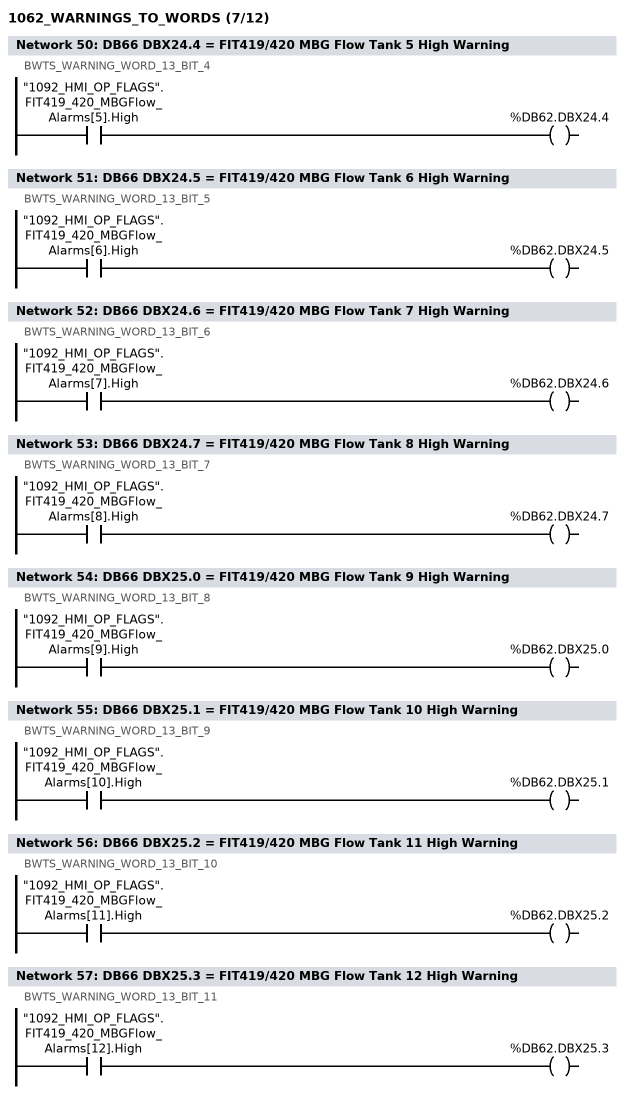
   RUNG wire#powerrail
      Contact( "1092_HMI_OP_FLAGS".FIT419_420_MBGFlow_Alarms[5].High )
      Coil( %DB62.DBX24.4 )
   END_RUNG
   // the same network as SCL:
   %DB62.DBX24.4 := "1092_HMI_OP_FLAGS".FIT419_420_MBGFlow_Alarms[5].High;
END_REGION

REGION Network 51: DB66 DBX24.5 = FIT419/420 MBG Flow Tank 6 High Warning
   // BWTS_WARNING_WORD_13_BIT_5
   RUNG wire#powerrail
      Contact( "1092_HMI_OP_FLAGS".FIT419_420_MBGFlow_Alarms[6].High )
      Coil( %DB62.DBX24.5 )
   END_RUNG
   // the same network as SCL:
   %DB62.DBX24.5 := "1092_HMI_OP_FLAGS".FIT419_420_MBGFlow_Alarms[6].High;
END_REGION

REGION Network 52: DB66 DBX24.6 = FIT419/420 MBG Flow Tank 7 High Warning
   // BWTS_WARNING_WORD_13_BIT_6
   RUNG wire#powerrail
      Contact( "1092_HMI_OP_FLAGS".FIT419_420_MBGFlow_Alarms[7].High )
      Coil( %DB62.DBX24.6 )
   END_RUNG
   // the same network as SCL:
   %DB62.DBX24.6 := "1092_HMI_OP_FLAGS".FIT419_420_MBGFlow_Alarms[7].High;
END_REGION

REGION Network 53: DB66 DBX24.7 = FIT419/420 MBG Flow Tank 8 High Warning
   // BWTS_WARNING_WORD_13_BIT_7
   RUNG wire#powerrail
      Contact( "1092_HMI_OP_FLAGS".FIT419_420_MBGFlow_Alarms[8].High )
      Coil( %DB62.DBX24.7 )
   END_RUNG
   // the same network as SCL:
   %DB62.DBX24.7 := "1092_HMI_OP_FLAGS".FIT419_420_MBGFlow_Alarms[8].High;
END_REGION

REGION Network 54: DB66 DBX25.0 = FIT419/420 MBG Flow Tank 9 High Warning
   // BWTS_WARNING_WORD_13_BIT_8
   RUNG wire#powerrail
      Contact( "1092_HMI_OP_FLAGS".FIT419_420_MBGFlow_Alarms[9].High )
      Coil( %DB62.DBX25.0 )
   END_RUNG
   // the same network as SCL:
   %DB62.DBX25.0 := "1092_HMI_OP_FLAGS".FIT419_420_MBGFlow_Alarms[9].High;
END_REGION

REGION Network 55: DB66 DBX25.1 = FIT419/420 MBG Flow Tank 10 High Warning
   // BWTS_WARNING_WORD_13_BIT_9
   RUNG wire#powerrail
      Contact( "1092_HMI_OP_FLAGS".FIT419_420_MBGFlow_Alarms[10].High )
      Coil( %DB62.DBX25.1 )
   END_RUNG
   // the same network as SCL:
   %DB62.DBX25.1 := "1092_HMI_OP_FLAGS".FIT419_420_MBGFlow_Alarms[10].High;
END_REGION

REGION Network 56: DB66 DBX25.2 = FIT419/420 MBG Flow Tank 11 High Warning
   // BWTS_WARNING_WORD_13_BIT_10
   RUNG wire#powerrail
      Contact( "1092_HMI_OP_FLAGS".FIT419_420_MBGFlow_Alarms[11].High )
      Coil( %DB62.DBX25.2 )
   END_RUNG
   // the same network as SCL:
   %DB62.DBX25.2 := "1092_HMI_OP_FLAGS".FIT419_420_MBGFlow_Alarms[11].High;
END_REGION

REGION Network 57: DB66 DBX25.3 = FIT419/420 MBG Flow Tank 12 High Warning
   // BWTS_WARNING_WORD_13_BIT_11
   RUNG wire#powerrail
      Contact( "1092_HMI_OP_FLAGS".FIT419_420_MBGFlow_Alarms[12].High )
      Coil( %DB62.DBX25.3 )
   END_RUNG
   // the same network as SCL:
   %DB62.DBX25.3 := "1092_HMI_OP_FLAGS".FIT419_420_MBGFlow_Alarms[12].High;
END_REGION

REGION Network 58: DB66 DBX25.4 = FIT419/420 MBG Flow Tank 13 High Warning
   // BWTS_WARNING_WORD_13_BIT_12
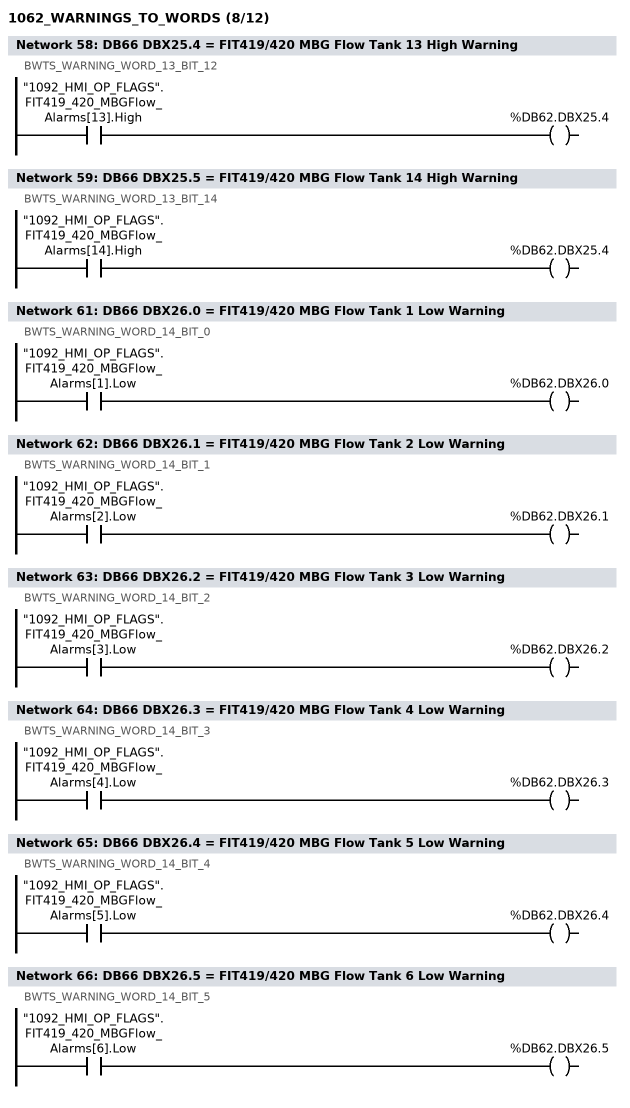
   RUNG wire#powerrail
      Contact( "1092_HMI_OP_FLAGS".FIT419_420_MBGFlow_Alarms[13].High )
      Coil( %DB62.DBX25.4 )
   END_RUNG
   // the same network as SCL:
   %DB62.DBX25.4 := "1092_HMI_OP_FLAGS".FIT419_420_MBGFlow_Alarms[13].High;
END_REGION

REGION Network 59: DB66 DBX25.5 = FIT419/420 MBG Flow Tank 14 High Warning
   // BWTS_WARNING_WORD_13_BIT_14
   RUNG wire#powerrail
      Contact( "1092_HMI_OP_FLAGS".FIT419_420_MBGFlow_Alarms[14].High )
      Coil( %DB62.DBX25.4 )
   END_RUNG
   // the same network as SCL:
   %DB62.DBX25.4 := "1092_HMI_OP_FLAGS".FIT419_420_MBGFlow_Alarms[14].High;
END_REGION

REGION Network 61: DB66 DBX26.0 = FIT419/420 MBG Flow Tank 1 Low Warning
   // BWTS_WARNING_WORD_14_BIT_0
   RUNG wire#powerrail
      Contact( "1092_HMI_OP_FLAGS".FIT419_420_MBGFlow_Alarms[1].Low )
      Coil( %DB62.DBX26.0 )
   END_RUNG
   // the same network as SCL:
   %DB62.DBX26.0 := "1092_HMI_OP_FLAGS".FIT419_420_MBGFlow_Alarms[1].Low;
END_REGION

REGION Network 62: DB66 DBX26.1 = FIT419/420 MBG Flow Tank 2 Low Warning
   // BWTS_WARNING_WORD_14_BIT_1
   RUNG wire#powerrail
      Contact( "1092_HMI_OP_FLAGS".FIT419_420_MBGFlow_Alarms[2].Low )
      Coil( %DB62.DBX26.1 )
   END_RUNG
   // the same network as SCL:
   %DB62.DBX26.1 := "1092_HMI_OP_FLAGS".FIT419_420_MBGFlow_Alarms[2].Low;
END_REGION

REGION Network 63: DB66 DBX26.2 = FIT419/420 MBG Flow Tank 3 Low Warning
   // BWTS_WARNING_WORD_14_BIT_2
   RUNG wire#powerrail
      Contact( "1092_HMI_OP_FLAGS".FIT419_420_MBGFlow_Alarms[3].Low )
      Coil( %DB62.DBX26.2 )
   END_RUNG
   // the same network as SCL:
   %DB62.DBX26.2 := "1092_HMI_OP_FLAGS".FIT419_420_MBGFlow_Alarms[3].Low;
END_REGION

REGION Network 64: DB66 DBX26.3 = FIT419/420 MBG Flow Tank 4 Low Warning
   // BWTS_WARNING_WORD_14_BIT_3
   RUNG wire#powerrail
      Contact( "1092_HMI_OP_FLAGS".FIT419_420_MBGFlow_Alarms[4].Low )
      Coil( %DB62.DBX26.3 )
   END_RUNG
   // the same network as SCL:
   %DB62.DBX26.3 := "1092_HMI_OP_FLAGS".FIT419_420_MBGFlow_Alarms[4].Low;
END_REGION

REGION Network 65: DB66 DBX26.4 = FIT419/420 MBG Flow Tank 5 Low Warning
   // BWTS_WARNING_WORD_14_BIT_4
   RUNG wire#powerrail
      Contact( "1092_HMI_OP_FLAGS".FIT419_420_MBGFlow_Alarms[5].Low )
      Coil( %DB62.DBX26.4 )
   END_RUNG
   // the same network as SCL:
   %DB62.DBX26.4 := "1092_HMI_OP_FLAGS".FIT419_420_MBGFlow_Alarms[5].Low;
END_REGION

REGION Network 66: DB66 DBX26.5 = FIT419/420 MBG Flow Tank 6 Low Warning
   // BWTS_WARNING_WORD_14_BIT_5
   RUNG wire#powerrail
      Contact( "1092_HMI_OP_FLAGS".FIT419_420_MBGFlow_Alarms[6].Low )
      Coil( %DB62.DBX26.5 )
   END_RUNG
   // the same network as SCL:
   %DB62.DBX26.5 := "1092_HMI_OP_FLAGS".FIT419_420_MBGFlow_Alarms[6].Low;
END_REGION

REGION Network 67: DB66 DBX26.6 = FIT419/420 MBG Flow Tank 7 Low Warning
   // BWTS_WARNING_WORD_14_BIT_6
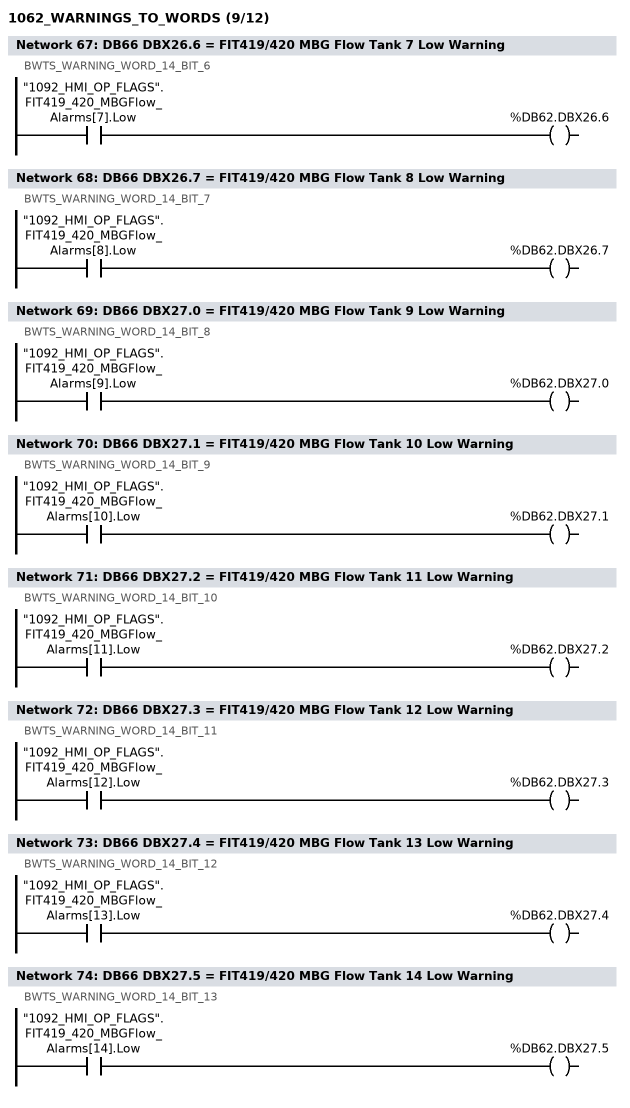
   RUNG wire#powerrail
      Contact( "1092_HMI_OP_FLAGS".FIT419_420_MBGFlow_Alarms[7].Low )
      Coil( %DB62.DBX26.6 )
   END_RUNG
   // the same network as SCL:
   %DB62.DBX26.6 := "1092_HMI_OP_FLAGS".FIT419_420_MBGFlow_Alarms[7].Low;
END_REGION

REGION Network 68: DB66 DBX26.7 = FIT419/420 MBG Flow Tank 8 Low Warning
   // BWTS_WARNING_WORD_14_BIT_7
   RUNG wire#powerrail
      Contact( "1092_HMI_OP_FLAGS".FIT419_420_MBGFlow_Alarms[8].Low )
      Coil( %DB62.DBX26.7 )
   END_RUNG
   // the same network as SCL:
   %DB62.DBX26.7 := "1092_HMI_OP_FLAGS".FIT419_420_MBGFlow_Alarms[8].Low;
END_REGION

REGION Network 69: DB66 DBX27.0 = FIT419/420 MBG Flow Tank 9 Low Warning
   // BWTS_WARNING_WORD_14_BIT_8
   RUNG wire#powerrail
      Contact( "1092_HMI_OP_FLAGS".FIT419_420_MBGFlow_Alarms[9].Low )
      Coil( %DB62.DBX27.0 )
   END_RUNG
   // the same network as SCL:
   %DB62.DBX27.0 := "1092_HMI_OP_FLAGS".FIT419_420_MBGFlow_Alarms[9].Low;
END_REGION

REGION Network 70: DB66 DBX27.1 = FIT419/420 MBG Flow Tank 10 Low Warning
   // BWTS_WARNING_WORD_14_BIT_9
   RUNG wire#powerrail
      Contact( "1092_HMI_OP_FLAGS".FIT419_420_MBGFlow_Alarms[10].Low )
      Coil( %DB62.DBX27.1 )
   END_RUNG
   // the same network as SCL:
   %DB62.DBX27.1 := "1092_HMI_OP_FLAGS".FIT419_420_MBGFlow_Alarms[10].Low;
END_REGION

REGION Network 71: DB66 DBX27.2 = FIT419/420 MBG Flow Tank 11 Low Warning
   // BWTS_WARNING_WORD_14_BIT_10
   RUNG wire#powerrail
      Contact( "1092_HMI_OP_FLAGS".FIT419_420_MBGFlow_Alarms[11].Low )
      Coil( %DB62.DBX27.2 )
   END_RUNG
   // the same network as SCL:
   %DB62.DBX27.2 := "1092_HMI_OP_FLAGS".FIT419_420_MBGFlow_Alarms[11].Low;
END_REGION

REGION Network 72: DB66 DBX27.3 = FIT419/420 MBG Flow Tank 12 Low Warning
   // BWTS_WARNING_WORD_14_BIT_11
   RUNG wire#powerrail
      Contact( "1092_HMI_OP_FLAGS".FIT419_420_MBGFlow_Alarms[12].Low )
      Coil( %DB62.DBX27.3 )
   END_RUNG
   // the same network as SCL:
   %DB62.DBX27.3 := "1092_HMI_OP_FLAGS".FIT419_420_MBGFlow_Alarms[12].Low;
END_REGION

REGION Network 73: DB66 DBX27.4 = FIT419/420 MBG Flow Tank 13 Low Warning
   // BWTS_WARNING_WORD_14_BIT_12
   RUNG wire#powerrail
      Contact( "1092_HMI_OP_FLAGS".FIT419_420_MBGFlow_Alarms[13].Low )
      Coil( %DB62.DBX27.4 )
   END_RUNG
   // the same network as SCL:
   %DB62.DBX27.4 := "1092_HMI_OP_FLAGS".FIT419_420_MBGFlow_Alarms[13].Low;
END_REGION

REGION Network 74: DB66 DBX27.5 = FIT419/420 MBG Flow Tank 14 Low Warning
   // BWTS_WARNING_WORD_14_BIT_13
   RUNG wire#powerrail
      Contact( "1092_HMI_OP_FLAGS".FIT419_420_MBGFlow_Alarms[14].Low )
      Coil( %DB62.DBX27.5 )
   END_RUNG
   // the same network as SCL:
   %DB62.DBX27.5 := "1092_HMI_OP_FLAGS".FIT419_420_MBGFlow_Alarms[14].Low;
END_REGION

REGION Network 76: DB66 DBX28.0 = PT424 Tank Group 1 High Warning
   // BWTS_WARNING_WORD_15_BIT_0
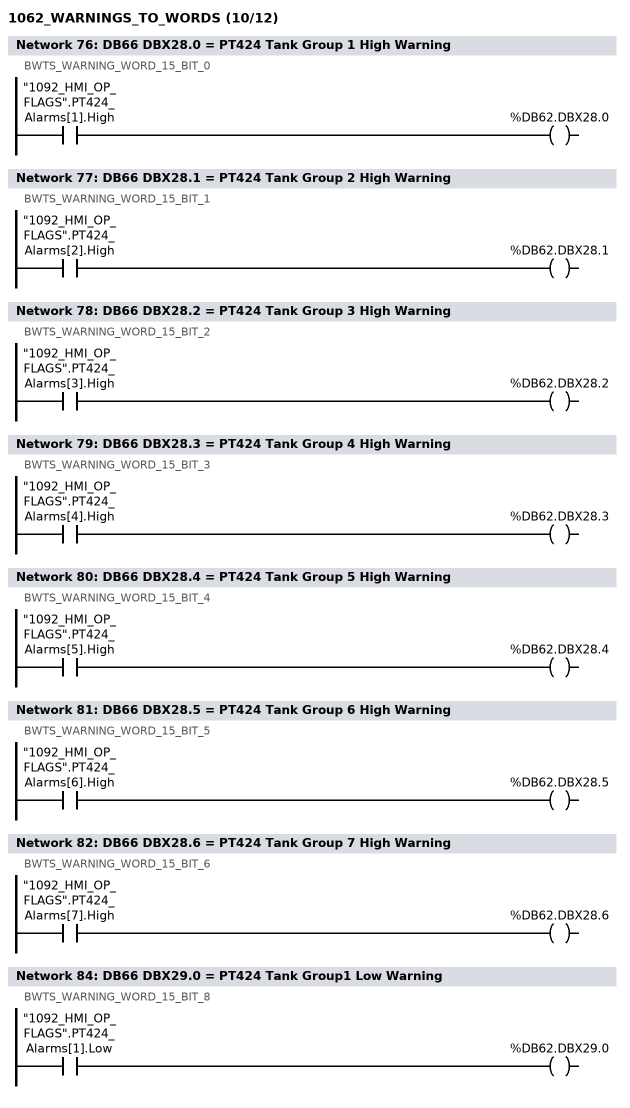
   RUNG wire#powerrail
      Contact( "1092_HMI_OP_FLAGS".PT424_Alarms[1].High )
      Coil( %DB62.DBX28.0 )
   END_RUNG
   // the same network as SCL:
   %DB62.DBX28.0 := "1092_HMI_OP_FLAGS".PT424_Alarms[1].High;
END_REGION

REGION Network 77: DB66 DBX28.1 = PT424 Tank Group 2 High Warning
   // BWTS_WARNING_WORD_15_BIT_1
   RUNG wire#powerrail
      Contact( "1092_HMI_OP_FLAGS".PT424_Alarms[2].High )
      Coil( %DB62.DBX28.1 )
   END_RUNG
   // the same network as SCL:
   %DB62.DBX28.1 := "1092_HMI_OP_FLAGS".PT424_Alarms[2].High;
END_REGION

REGION Network 78: DB66 DBX28.2 = PT424 Tank Group 3 High Warning
   // BWTS_WARNING_WORD_15_BIT_2
   RUNG wire#powerrail
      Contact( "1092_HMI_OP_FLAGS".PT424_Alarms[3].High )
      Coil( %DB62.DBX28.2 )
   END_RUNG
   // the same network as SCL:
   %DB62.DBX28.2 := "1092_HMI_OP_FLAGS".PT424_Alarms[3].High;
END_REGION

REGION Network 79: DB66 DBX28.3 = PT424 Tank Group 4 High Warning
   // BWTS_WARNING_WORD_15_BIT_3
   RUNG wire#powerrail
      Contact( "1092_HMI_OP_FLAGS".PT424_Alarms[4].High )
      Coil( %DB62.DBX28.3 )
   END_RUNG
   // the same network as SCL:
   %DB62.DBX28.3 := "1092_HMI_OP_FLAGS".PT424_Alarms[4].High;
END_REGION

REGION Network 80: DB66 DBX28.4 = PT424 Tank Group 5 High Warning
   // BWTS_WARNING_WORD_15_BIT_4
   RUNG wire#powerrail
      Contact( "1092_HMI_OP_FLAGS".PT424_Alarms[5].High )
      Coil( %DB62.DBX28.4 )
   END_RUNG
   // the same network as SCL:
   %DB62.DBX28.4 := "1092_HMI_OP_FLAGS".PT424_Alarms[5].High;
END_REGION

REGION Network 81: DB66 DBX28.5 = PT424 Tank Group 6 High Warning
   // BWTS_WARNING_WORD_15_BIT_5
   RUNG wire#powerrail
      Contact( "1092_HMI_OP_FLAGS".PT424_Alarms[6].High )
      Coil( %DB62.DBX28.5 )
   END_RUNG
   // the same network as SCL:
   %DB62.DBX28.5 := "1092_HMI_OP_FLAGS".PT424_Alarms[6].High;
END_REGION

REGION Network 82: DB66 DBX28.6 = PT424 Tank Group 7 High Warning
   // BWTS_WARNING_WORD_15_BIT_6
   RUNG wire#powerrail
      Contact( "1092_HMI_OP_FLAGS".PT424_Alarms[7].High )
      Coil( %DB62.DBX28.6 )
   END_RUNG
   // the same network as SCL:
   %DB62.DBX28.6 := "1092_HMI_OP_FLAGS".PT424_Alarms[7].High;
END_REGION

REGION Network 84: DB66 DBX29.0 = PT424 Tank Group1 Low Warning
   // BWTS_WARNING_WORD_15_BIT_8
   RUNG wire#powerrail
      Contact( "1092_HMI_OP_FLAGS".PT424_Alarms[1].Low )
      Coil( %DB62.DBX29.0 )
   END_RUNG
   // the same network as SCL:
   %DB62.DBX29.0 := "1092_HMI_OP_FLAGS".PT424_Alarms[1].Low;
END_REGION

REGION Network 85: DB66 DBX29.1 = PT424 Tank Group 2 Low Warning
   // BWTS_WARNING_WORD_15_BIT_9
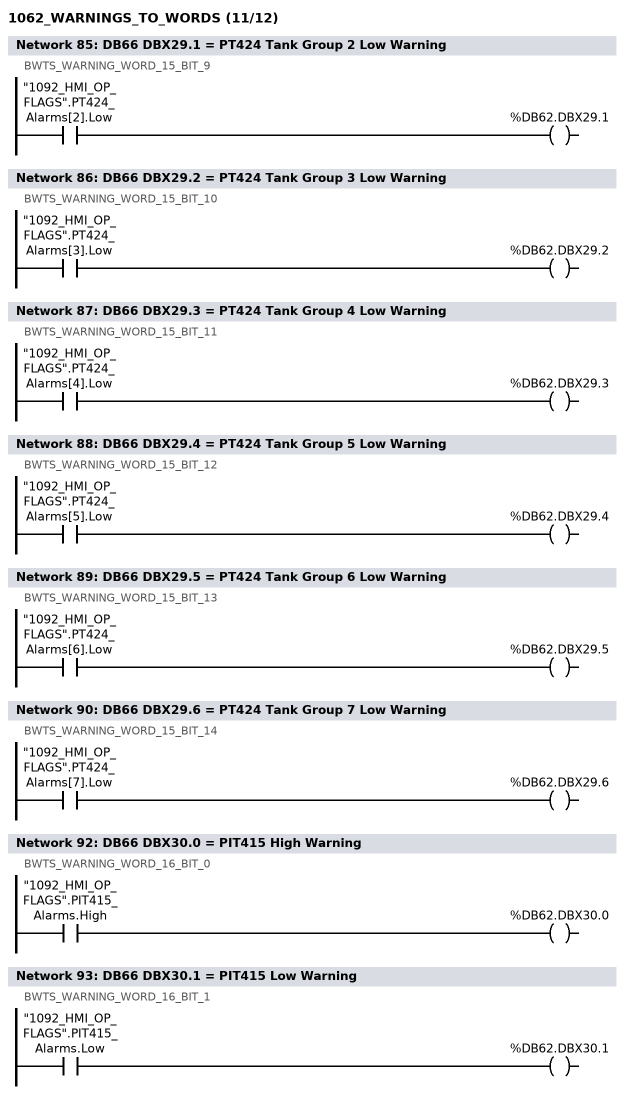
   RUNG wire#powerrail
      Contact( "1092_HMI_OP_FLAGS".PT424_Alarms[2].Low )
      Coil( %DB62.DBX29.1 )
   END_RUNG
   // the same network as SCL:
   %DB62.DBX29.1 := "1092_HMI_OP_FLAGS".PT424_Alarms[2].Low;
END_REGION

REGION Network 86: DB66 DBX29.2 = PT424 Tank Group 3 Low Warning
   // BWTS_WARNING_WORD_15_BIT_10
   RUNG wire#powerrail
      Contact( "1092_HMI_OP_FLAGS".PT424_Alarms[3].Low )
      Coil( %DB62.DBX29.2 )
   END_RUNG
   // the same network as SCL:
   %DB62.DBX29.2 := "1092_HMI_OP_FLAGS".PT424_Alarms[3].Low;
END_REGION

REGION Network 87: DB66 DBX29.3 = PT424 Tank Group 4 Low Warning
   // BWTS_WARNING_WORD_15_BIT_11
   RUNG wire#powerrail
      Contact( "1092_HMI_OP_FLAGS".PT424_Alarms[4].Low )
      Coil( %DB62.DBX29.3 )
   END_RUNG
   // the same network as SCL:
   %DB62.DBX29.3 := "1092_HMI_OP_FLAGS".PT424_Alarms[4].Low;
END_REGION

REGION Network 88: DB66 DBX29.4 = PT424 Tank Group 5 Low Warning
   // BWTS_WARNING_WORD_15_BIT_12
   RUNG wire#powerrail
      Contact( "1092_HMI_OP_FLAGS".PT424_Alarms[5].Low )
      Coil( %DB62.DBX29.4 )
   END_RUNG
   // the same network as SCL:
   %DB62.DBX29.4 := "1092_HMI_OP_FLAGS".PT424_Alarms[5].Low;
END_REGION

REGION Network 89: DB66 DBX29.5 = PT424 Tank Group 6 Low Warning
   // BWTS_WARNING_WORD_15_BIT_13
   RUNG wire#powerrail
      Contact( "1092_HMI_OP_FLAGS".PT424_Alarms[6].Low )
      Coil( %DB62.DBX29.5 )
   END_RUNG
   // the same network as SCL:
   %DB62.DBX29.5 := "1092_HMI_OP_FLAGS".PT424_Alarms[6].Low;
END_REGION

REGION Network 90: DB66 DBX29.6 = PT424 Tank Group 7 Low Warning
   // BWTS_WARNING_WORD_15_BIT_14
   RUNG wire#powerrail
      Contact( "1092_HMI_OP_FLAGS".PT424_Alarms[7].Low )
      Coil( %DB62.DBX29.6 )
   END_RUNG
   // the same network as SCL:
   %DB62.DBX29.6 := "1092_HMI_OP_FLAGS".PT424_Alarms[7].Low;
END_REGION

REGION Network 92: DB66 DBX30.0 = PIT415 High Warning
   // BWTS_WARNING_WORD_16_BIT_0
   RUNG wire#powerrail
      Contact( "1092_HMI_OP_FLAGS".PIT415_Alarms.High )
      Coil( %DB62.DBX30.0 )
   END_RUNG
   // the same network as SCL:
   %DB62.DBX30.0 := "1092_HMI_OP_FLAGS".PIT415_Alarms.High;
END_REGION

REGION Network 93: DB66 DBX30.1 = PIT415 Low Warning
   // BWTS_WARNING_WORD_16_BIT_1
   RUNG wire#powerrail
      Contact( "1092_HMI_OP_FLAGS".PIT415_Alarms.Low )
      Coil( %DB62.DBX30.1 )
   END_RUNG
   // the same network as SCL:
   %DB62.DBX30.1 := "1092_HMI_OP_FLAGS".PIT415_Alarms.Low;
END_REGION

REGION Network 95: Warning Present
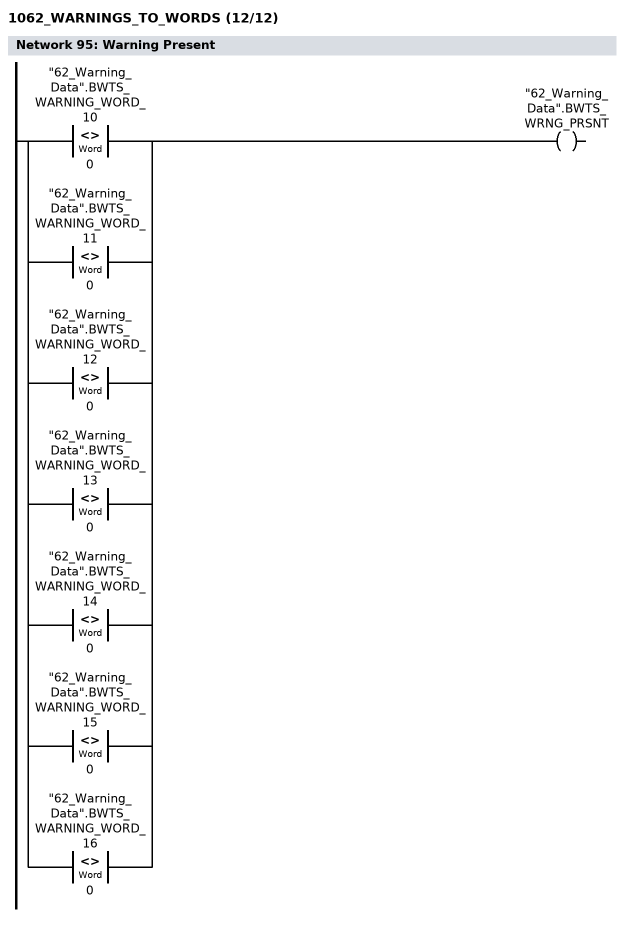
   RUNG wire#powerrail
      { S7_Templates := "SrcType := Word" } NE_Contact(in1 := "62_Warning_Data".BWTS_WARNING_WORD_10, in2 := 0)
      wire#w1
      Coil( "62_Warning_Data".BWTS_WRNG_PRSNT )
   END_RUNG
   RUNG wire#powerrail
      { S7_Templates := "SrcType := Word" } NE_Contact(in1 := "62_Warning_Data".BWTS_WARNING_WORD_11, in2 := 0)
   END_RUNG wire#w1
   RUNG wire#powerrail
      { S7_Templates := "SrcType := Word" } NE_Contact(in1 := "62_Warning_Data".BWTS_WARNING_WORD_12, in2 := 0)
   END_RUNG wire#w1
   RUNG wire#powerrail
      { S7_Templates := "SrcType := Word" } NE_Contact(in1 := "62_Warning_Data".BWTS_WARNING_WORD_13, in2 := 0)
   END_RUNG wire#w1
   RUNG wire#powerrail
      { S7_Templates := "SrcType := Word" } NE_Contact(in1 := "62_Warning_Data".BWTS_WARNING_WORD_14, in2 := 0)
   END_RUNG wire#w1
   RUNG wire#powerrail
      { S7_Templates := "SrcType := Word" } NE_Contact(in1 := "62_Warning_Data".BWTS_WARNING_WORD_15, in2 := 0)
   END_RUNG wire#w1
   RUNG wire#powerrail
      { S7_Templates := "SrcType := Word" } NE_Contact(in1 := "62_Warning_Data".BWTS_WARNING_WORD_16, in2 := 0)
   END_RUNG wire#w1
   // the same network as SCL:
   "62_Warning_Data".BWTS_WRNG_PRSNT := ("62_Warning_Data".BWTS_WARNING_WORD_10 <> 0) OR ("62_Warning_Data".BWTS_WARNING_WORD_11 <> 0) OR ("62_Warning_Data".BWTS_WARNING_WORD_12 <> 0) OR ("62_Warning_Data".BWTS_WARNING_WORD_13 <> 0) OR ("62_Warning_Data".BWTS_WARNING_WORD_14 <> 0) OR ("62_Warning_Data".BWTS_WARNING_WORD_15 <> 0) OR ("62_Warning_Data".BWTS_WARNING_WORD_16 <> 0);
END_REGION
END_FUNCTION

FUNCTION "1065_MANAGE_ONEOFF_ALARMS" : Void   // FC1065, LAD
{ S7_Optimized_Access := 'TRUE' }
VERSION : 0.1
// Manage all one-off alarms that do not assign to a tank or tank group directly.
// Note: This function calls analog health trips directly.
   VAR_TEMP
      DummyAlarm : Bool;
   END_VAR
BEGIN

REGION Network 1: PIT415 (Deck Main IG) Alarm
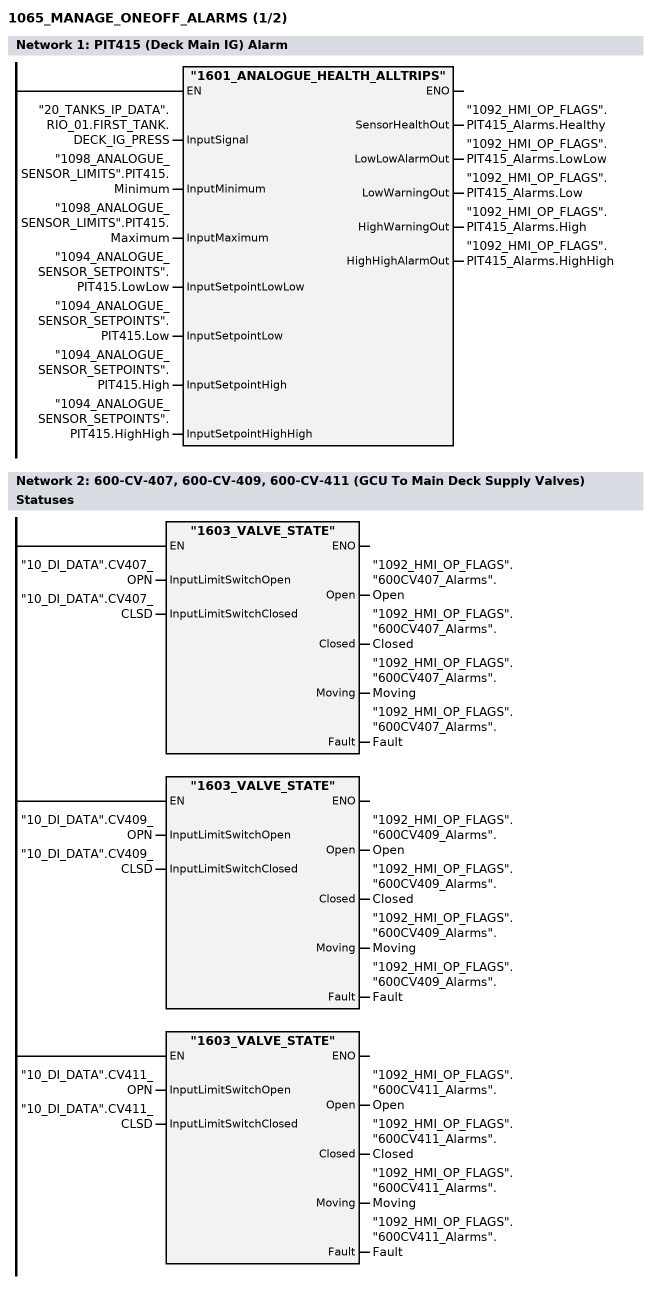
   RUNG wire#powerrail
      "1601_ANALOGUE_HEALTH_ALLTRIPS"(InputSignal := "20_TANKS_IP_DATA".RIO_01.FIRST_TANK.DECK_IG_PRESS, InputMinimum := "1098_ANALOGUE_SENSOR_LIMITS".PIT415.Minimum, InputMaximum := "1098_ANALOGUE_SENSOR_LIMITS".PIT415.Maximum, InputSetpointLowLow := "1094_ANALOGUE_SENSOR_SETPOINTS".PIT415.LowLow, InputSetpointLow := "1094_ANALOGUE_SENSOR_SETPOINTS".PIT415.Low, InputSetpointHigh := "1094_ANALOGUE_SENSOR_SETPOINTS".PIT415.High, InputSetpointHighHigh := "1094_ANALOGUE_SENSOR_SETPOINTS".PIT415.HighHigh, SensorHealthOut => "1092_HMI_OP_FLAGS".PIT415_Alarms.Healthy, LowLowAlarmOut => "1092_HMI_OP_FLAGS".PIT415_Alarms.LowLow, LowWarningOut => "1092_HMI_OP_FLAGS".PIT415_Alarms.Low, HighWarningOut => "1092_HMI_OP_FLAGS".PIT415_Alarms.High, HighHighAlarmOut => "1092_HMI_OP_FLAGS".PIT415_Alarms.HighHigh)
   END_RUNG
   // the same network as SCL:
   "1601_ANALOGUE_HEALTH_ALLTRIPS"(InputSignal := "20_TANKS_IP_DATA".RIO_01.FIRST_TANK.DECK_IG_PRESS,
                           InputMinimum := "1098_ANALOGUE_SENSOR_LIMITS".PIT415.Minimum,
                           InputMaximum := "1098_ANALOGUE_SENSOR_LIMITS".PIT415.Maximum,
                           InputSetpointLowLow := "1094_ANALOGUE_SENSOR_SETPOINTS".PIT415.LowLow,
                           InputSetpointLow := "1094_ANALOGUE_SENSOR_SETPOINTS".PIT415.Low,
                           InputSetpointHigh := "1094_ANALOGUE_SENSOR_SETPOINTS".PIT415.High,
                           InputSetpointHighHigh := "1094_ANALOGUE_SENSOR_SETPOINTS".PIT415.HighHigh,
                           SensorHealthOut => "1092_HMI_OP_FLAGS".PIT415_Alarms.Healthy,
                           LowLowAlarmOut => "1092_HMI_OP_FLAGS".PIT415_Alarms.LowLow,
                           LowWarningOut => "1092_HMI_OP_FLAGS".PIT415_Alarms.Low,
                           HighWarningOut => "1092_HMI_OP_FLAGS".PIT415_Alarms.High,
                           HighHighAlarmOut => "1092_HMI_OP_FLAGS".PIT415_Alarms.HighHigh);
END_REGION

REGION Network 2: 600-CV-407, 600-CV-409, 600-CV-411 (GCU To Main Deck Supply Valves) Statuses
   RUNG wire#powerrail
      "1603_VALVE_STATE"(InputLimitSwitchOpen := "10_DI_DATA".CV407_OPN, InputLimitSwitchClosed := "10_DI_DATA".CV407_CLSD, Open => "1092_HMI_OP_FLAGS"."600CV407_Alarms".Open, Closed => "1092_HMI_OP_FLAGS"."600CV407_Alarms".Closed, Moving => "1092_HMI_OP_FLAGS"."600CV407_Alarms".Moving, Fault => "1092_HMI_OP_FLAGS"."600CV407_Alarms".Fault)
   END_RUNG
   RUNG wire#powerrail
      "1603_VALVE_STATE"(InputLimitSwitchOpen := "10_DI_DATA".CV409_OPN, InputLimitSwitchClosed := "10_DI_DATA".CV409_CLSD, Open => "1092_HMI_OP_FLAGS"."600CV409_Alarms".Open, Closed => "1092_HMI_OP_FLAGS"."600CV409_Alarms".Closed, Moving => "1092_HMI_OP_FLAGS"."600CV409_Alarms".Moving, Fault => "1092_HMI_OP_FLAGS"."600CV409_Alarms".Fault)
   END_RUNG
   RUNG wire#powerrail
      "1603_VALVE_STATE"(InputLimitSwitchOpen := "10_DI_DATA".CV411_OPN, InputLimitSwitchClosed := "10_DI_DATA".CV411_CLSD, Open => "1092_HMI_OP_FLAGS"."600CV411_Alarms".Open, Closed => "1092_HMI_OP_FLAGS"."600CV411_Alarms".Closed, Moving => "1092_HMI_OP_FLAGS"."600CV411_Alarms".Moving, Fault => "1092_HMI_OP_FLAGS"."600CV411_Alarms".Fault)
   END_RUNG
   // the same network as SCL:
   "1603_VALVE_STATE"(InputLimitSwitchOpen := "10_DI_DATA".CV407_OPN,
                      InputLimitSwitchClosed := "10_DI_DATA".CV407_CLSD,
                      Open => "1092_HMI_OP_FLAGS"."600CV407_Alarms".Open,
                      Closed => "1092_HMI_OP_FLAGS"."600CV407_Alarms".Closed,
                      Moving => "1092_HMI_OP_FLAGS"."600CV407_Alarms".Moving,
                      Fault => "1092_HMI_OP_FLAGS"."600CV407_Alarms".Fault);
   "1603_VALVE_STATE"(InputLimitSwitchOpen := "10_DI_DATA".CV409_OPN,
                      InputLimitSwitchClosed := "10_DI_DATA".CV409_CLSD,
                      Open => "1092_HMI_OP_FLAGS"."600CV409_Alarms".Open,
                      Closed => "1092_HMI_OP_FLAGS"."600CV409_Alarms".Closed,
                      Moving => "1092_HMI_OP_FLAGS"."600CV409_Alarms".Moving,
                      Fault => "1092_HMI_OP_FLAGS"."600CV409_Alarms".Fault);
   "1603_VALVE_STATE"(InputLimitSwitchOpen := "10_DI_DATA".CV411_OPN,
                      InputLimitSwitchClosed := "10_DI_DATA".CV411_CLSD,
                      Open => "1092_HMI_OP_FLAGS"."600CV411_Alarms".Open,
                      Closed => "1092_HMI_OP_FLAGS"."600CV411_Alarms".Closed,
                      Moving => "1092_HMI_OP_FLAGS"."600CV411_Alarms".Moving,
                      Fault => "1092_HMI_OP_FLAGS"."600CV411_Alarms".Fault);
END_REGION

REGION Network 3: TX-430 (Salinometer) Alarm
   // Note: This block does not apply to any requirments in BWTS as of 20/02/2019, but has been communicated via e-mail from CHM to FNC. The salinometer has previously been called SL400.
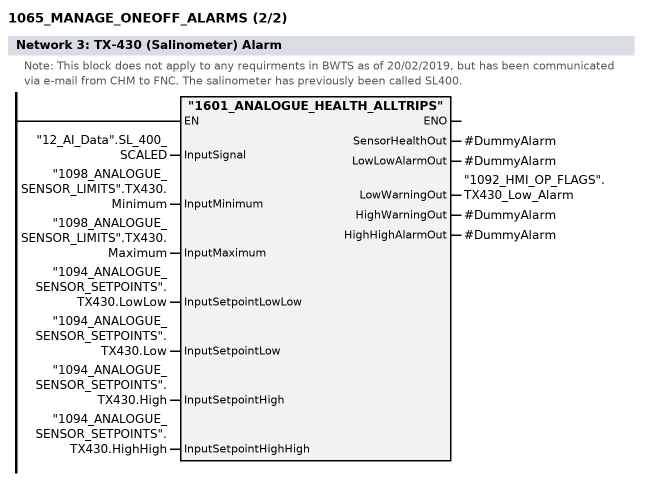
   RUNG wire#powerrail
      "1601_ANALOGUE_HEALTH_ALLTRIPS"(InputSignal := "12_AI_Data".SL_400_SCALED, InputMinimum := "1098_ANALOGUE_SENSOR_LIMITS".TX430.Minimum, InputMaximum := "1098_ANALOGUE_SENSOR_LIMITS".TX430.Maximum, InputSetpointLowLow := "1094_ANALOGUE_SENSOR_SETPOINTS".TX430.LowLow, InputSetpointLow := "1094_ANALOGUE_SENSOR_SETPOINTS".TX430.Low, InputSetpointHigh := "1094_ANALOGUE_SENSOR_SETPOINTS".TX430.High, InputSetpointHighHigh := "1094_ANALOGUE_SENSOR_SETPOINTS".TX430.HighHigh, SensorHealthOut => #DummyAlarm, LowLowAlarmOut => #DummyAlarm, LowWarningOut => "1092_HMI_OP_FLAGS".TX430_Low_Alarm, HighWarningOut => #DummyAlarm, HighHighAlarmOut => #DummyAlarm)
   END_RUNG
   // the same network as SCL:
   "1601_ANALOGUE_HEALTH_ALLTRIPS"(InputSignal := "12_AI_Data".SL_400_SCALED,
                           InputMinimum := "1098_ANALOGUE_SENSOR_LIMITS".TX430.Minimum,
                           InputMaximum := "1098_ANALOGUE_SENSOR_LIMITS".TX430.Maximum,
                           InputSetpointLowLow := "1094_ANALOGUE_SENSOR_SETPOINTS".TX430.LowLow,
                           InputSetpointLow := "1094_ANALOGUE_SENSOR_SETPOINTS".TX430.Low,
                           InputSetpointHigh := "1094_ANALOGUE_SENSOR_SETPOINTS".TX430.High,
                           InputSetpointHighHigh := "1094_ANALOGUE_SENSOR_SETPOINTS".TX430.HighHigh,
                           SensorHealthOut => #DummyAlarm,
                           LowLowAlarmOut => #DummyAlarm,
                           LowWarningOut => "1092_HMI_OP_FLAGS".TX430_Low_Alarm,
                           HighWarningOut => #DummyAlarm,
                           HighHighAlarmOut => #DummyAlarm);
END_REGION
END_FUNCTION

FUNCTION "1066_MANAGE_TANK_ALARMS" : Void   // FC1066, LAD
{ S7_Optimized_Access := 'TRUE' }
VERSION : 0.1
// Manage all alarms which are related to each tank (one alarm set per tank).
// Note: This function calls a wrapper for each sensor type which contains the alarm calculations.
// Note: TX427 and TX428 alarms use differing setpoints based on the phase of the system, see sub-function for futher information.
BEGIN

REGION Network 1: LT421, LT422 (BWTLevel) Alarms (All)
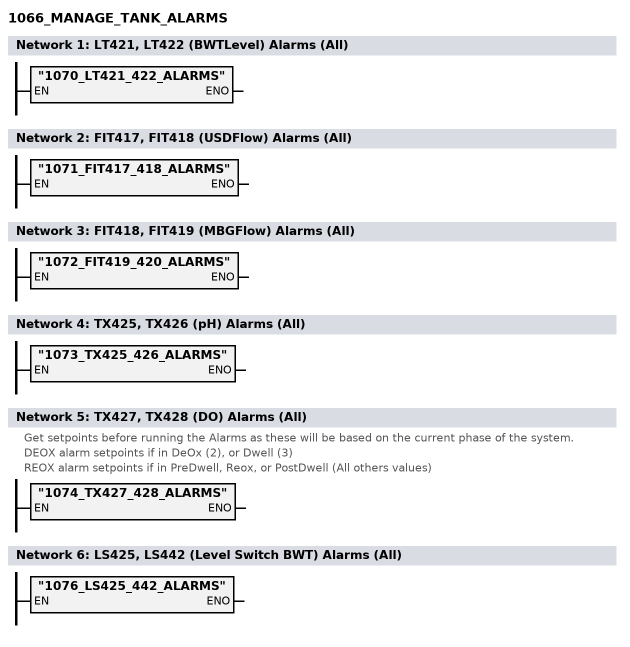
   RUNG wire#powerrail
      "1070_LT421_422_ALARMS"()
   END_RUNG
   // the same network as SCL:
   "1070_LT421_422_ALARMS"();
END_REGION

REGION Network 2: FIT417, FIT418 (USDFlow) Alarms (All)
   RUNG wire#powerrail
      "1071_FIT417_418_ALARMS"()
   END_RUNG
   // the same network as SCL:
   "1071_FIT417_418_ALARMS"();
END_REGION

REGION Network 3: FIT418, FIT419 (MBGFlow) Alarms (All)
   RUNG wire#powerrail
      "1072_FIT419_420_ALARMS"()
   END_RUNG
   // the same network as SCL:
   "1072_FIT419_420_ALARMS"();
END_REGION

REGION Network 4: TX425, TX426 (pH) Alarms (All)
   RUNG wire#powerrail
      "1073_TX425_426_ALARMS"()
   END_RUNG
   // the same network as SCL:
   "1073_TX425_426_ALARMS"();
END_REGION

REGION Network 5: TX427, TX428 (DO) Alarms (All)
   // Get setpoints before running the Alarms as these will be based on the current phase of the system.
   //     DEOX alarm setpoints if in DeOx (2), or Dwell (3)
   //     REOX alarm setpoints if in PreDwell, Reox, or PostDwell (All others values)
   RUNG wire#powerrail
      "1074_TX427_428_ALARMS"()
   END_RUNG
   // the same network as SCL:
   "1074_TX427_428_ALARMS"();
END_REGION

REGION Network 6: LS425, LS442 (Level Switch BWT) Alarms (All)
   RUNG wire#powerrail
      "1076_LS425_442_ALARMS"()
   END_RUNG
   // the same network as SCL:
   "1076_LS425_442_ALARMS"();
END_REGION
END_FUNCTION

FUNCTION "1067_MANAGE_TANKGROUP_ALARMS" : Void   // FC1067, LAD
{ S7_Optimized_Access := 'TRUE' }
VERSION : 0.1
// Manage all alarms which are related to a tank group (one alarm set per tank group).
// Note: This function calls a wrapper for each sensor type which contains the alarm calculations.
BEGIN

REGION Network 1: PT424 Alarms (Ullage Space Pressure Transmitter) (All)
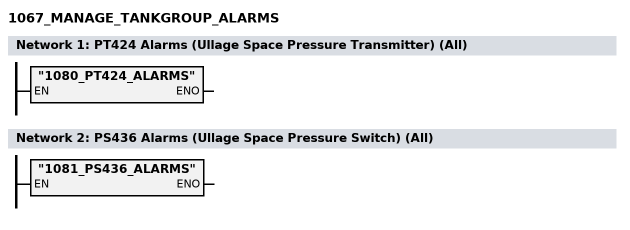
   RUNG wire#powerrail
      "1080_PT424_ALARMS"()
   END_RUNG
   // the same network as SCL:
   "1080_PT424_ALARMS"();
END_REGION

REGION Network 2: PS436 Alarms (Ullage Space Pressure Switch) (All)
   RUNG wire#powerrail
      "1081_PS436_ALARMS"()
   END_RUNG
   // the same network as SCL:
   "1081_PS436_ALARMS"();
END_REGION
END_FUNCTION

FUNCTION "1068_MANAGE_VALVE_STATUS" : Void   // FC1068, LAD
{ S7_Optimized_Access := 'TRUE' }
VERSION : 0.1
// Manage all valve position status'.
// Note: This function calls a wrapper for each valve type which contains the valve calculations.
// Note: If pressure valves are used in this system the alarms are not reported for PVVA/B valves and are suppressed here.
BEGIN

REGION Network 1: 600-CV-421, 600-CV-422 (Gas To Tank Inlet Valves) Statuses (All)